// TIA Portal project "N16-1166-5_27082020" (V13)

(* hardware
DEVICE "S71500/ET200MP station_1"  S7-1500 station
   slot 0: "Rail_0"  6ES7 590-1***0-0AA0
   slot 1: "PLC1"  CPU 1513-1 PN  6ES7 513-1AL01-0AB0  V1.8
DEVICE "ET 200SP station_1"  ET 200SP-Station
   slot 0: "Rack_0"  6ES5 710-8MAx1
   slot 0: "pa30"  IM155-6 PN BA  6ES7 155-6AR00-0AN0  V3.2
   slot 1: "DI A11"  DI 8x24VDC ST  6ES7 131-6BF00-0BA0  V1.1
      slot 1: "DI A11"  DI 8x24VDC ST  6ES7 131-6BF00-0BA0
   slot 2: "DI A12"  DI 8x24VDC ST  6ES7 131-6BF00-0BA0  V1.0
      slot 1: "DI A12"  DI 8x24VDC ST  6ES7 131-6BF00-0BA0
   slot 3: "DQ A13"  8DO 24VDC/0,5A ST  6ES7 132-6BF00-0BA0  V1.1
      slot 1: "DQ A13"  DQ 8x24VDC/0.5A ST  6ES7 132-6BF00-0BA0
   slot 4: "CM PtP A14"  CM PtP  6ES7 137-6AA00-0BA0  V1.0
      slot 1: "CM PtP A14"  CM PtP Sub  6ES7 137-6AA00-0BA0
   slot 5: "DI A15"  DI 16x24VDC ST  6ES7 131-6BH00-0BA0  V1.1
      slot 1: "DI A15"  DI 16x24VDC ST  6ES7 131-6BH00-0BA0
   slot 6: "DQ A16"  DQ 16x24VDC/0.5A ST  6ES7 132-6BH00-0BA0  V1.1
      slot 1: "DQ A16"  DQ 16x24VDC/0.5A ST  6ES7 132-6BH00-0BA0
   slot 7: "DI A17"  DI 8x24VDC ST  6ES7 131-6BF00-0BA0  V1.1
      slot 1: "DI A17"  DI 8x24VDC ST  6ES7 131-6BF00-0BA0
   slot 8: "Server module_1"  Server module  6ES7 193-6PA00-0AA0  V1.0
      slot 1: "Server module_1"  Server module  6ES7 193-6PA00-0AA0
   slot 127: "PROFINET BusAdapter CU"  PROFINET Interface  6ES7 193-6AR00-0AA0  V0.0
      slot 1: "Port_1"  6ES7 193-6AR00-0AA0  V0.0
      slot 2: "Port_2"  6ES7 193-6AR00-0AA0  V0.0
DEVICE "ET 200SP station_3"  ET 200SP-Station
   slot 0: "Rack_0"  6ES5 710-8MAx1
   slot 0: "pa60"  IM155-6 PN BA  6ES7 155-6AR00-0AN0  V3.2
   slot 1: "DI 8x24VDC ST_1"  DI 8x24VDC ST  6ES7 131-6BF00-0BA0  V1.1
      slot 1: "DI 8x24VDC ST_1"  DI 8x24VDC ST  6ES7 131-6BF00-0BA0
   slot 2: "DI 8x24VDC ST_2"  DI 8x24VDC ST  6ES7 131-6BF00-0BA0  V1.0
      slot 1: "DI 8x24VDC ST_2"  DI 8x24VDC ST  6ES7 131-6BF00-0BA0
   slot 3: "DI 8x24VDC ST_3"  DI 8x24VDC ST  6ES7 131-6BF00-0BA0  V1.1
      slot 1: "DI 8x24VDC ST_3"  DI 8x24VDC ST  6ES7 131-6BF00-0BA0
   slot 4: "DQ 8x24VDC/0.5A ST_1"  8DO 24VDC/0,5A ST  6ES7 132-6BF00-0BA0  V1.1
      slot 1: "DQ 8x24VDC/0.5A ST_1"  DQ 8x24VDC/0.5A ST  6ES7 132-6BF00-0BA0
   slot 5: "CM PtP_1"  CM PtP  6ES7 137-6AA00-0BA0  V1.0
      slot 1: "CM PtP_1"  CM PtP Sub  6ES7 137-6AA00-0BA0
   slot 6: "DI 16x24VDC ST_1"  DI 16x24VDC ST  6ES7 131-6BH00-0BA0  V1.1
      slot 1: "DI 16x24VDC ST_1"  DI 16x24VDC ST  6ES7 131-6BH00-0BA0
   slot 7: "DQ 16x24VDC/0.5A ST_1"  DQ 16x24VDC/0.5A ST  6ES7 132-6BH00-0BA0  V1.1
      slot 1: "DQ 16x24VDC/0.5A ST_1"  DQ 16x24VDC/0.5A ST  6ES7 132-6BH00-0BA0
   slot 8: "Server module_1"  Server module  6ES7 193-6PA00-0AA0  V1.0
      slot 1: "Server module_1"  Server module  6ES7 193-6PA00-0AA0
   slot 127: "PROFINET BusAdapter CU"  PROFINET Interface  6ES7 193-6AR00-0AA0  V0.0
      slot 1: "Port_1"  6ES7 193-6AR00-0AA0  V0.0
      slot 2: "Port_2"  6ES7 193-6AR00-0AA0  V0.0
DEVICE "HMI_pa30"  KTP700 Basic PN
   slot 0: "HMI"  HMI  6AV2 123-2GB03-0AX0  13.0.1.0
   slot 1: "HMI_RT_2"  KTP700 Basic PN  6AV2 123-2GB03-0AX0  13.0.1.0
   slot 5: "HMI_pa30.IE_CP_1"  PROFINET Interface
      slot 1: "PROFINET Interface_1"  PROFINET Interface
         slot 1: "Port_1"  Port
DEVICE "HMI_pa60"  KTP700 Basic PN
   slot 0: "HMI"  HMI  6AV2 123-2GB03-0AX0  13.0.1.0
   slot 1: "HMI_RT_4"  KTP700 Basic PN  6AV2 123-2GB03-0AX0  13.0.1.0
   slot 5: "HMI_pa60.IE_CP_1"  PROFINET Interface
      slot 1: "PROFINET Interface_1"  PROFINET Interface
         slot 1: "Port_1"  Port
DEVICE "ET 200SP station_4"  ET 200SP-Station
   slot 0: "Rack_0"  6ES5 710-8MAx1
   slot 0: "LightControll"  IM155-6 PN BA  6ES7 155-6AR00-0AN0  V3.2
   slot 1: "DQ 16x24VDC/0.5A ST_1"  DQ 16x24VDC/0.5A ST  6ES7 132-6BH00-0BA0  V1.1
      slot 1: "DQ 16x24VDC/0.5A ST_1"  DQ 16x24VDC/0.5A ST  6ES7 132-6BH00-0BA0
   slot 2: "Server module_1"  Server module  6ES7 193-6PA00-0AA0  V1.0
      slot 1: "Server module_1"  Server module  6ES7 193-6PA00-0AA0
   slot 127: "PROFINET BusAdapter CU"  PROFINET Interface  6ES7 193-6AR00-0AA0  V0.0
      slot 1: "Port_1"  6ES7 193-6AR00-0AA0  V0.0
      slot 2: "Port_2"  6ES7 193-6AR00-0AA0  V0.0
DEVICE "S71500/ET200MP station_2"  S7-1500 station
   slot 0: "Rail_0"  6ES7 590-1***0-0AA0
   slot 2: "CP 1543-1_1"  CP 1543-1  6GK7 543-1AX00-0XE0  V1.1
DEVICE "HMI_PA10B"  KTP700 Basic PN
   slot 0: "HMI"  HMI  6AV2 123-2GB03-0AX0  13.0.1.0
   slot 1: "HMI_RT_5"  KTP700 Basic PN  6AV2 123-2GB03-0AX0  13.0.1.0
   slot 5: "HMI_PA10B.IE_CP_1"  PROFINET Interface
      slot 1: "PROFINET Interface_1"  PROFINET Interface
         slot 1: "Port_1"  Port
DEVICE "ET 200SP station_5"  ET 200SP-Station
   slot 0: "Rack_0"  6ES5 710-8MAx1
   slot 0: "FS"  IM155-6 PN BA  6ES7 155-6AR00-0AN0  V3.2
   slot 1: "DI 8x24VDC ST_1"  DI 8x24VDC ST  6ES7 131-6BF00-0BA0  V1.0
      slot 1: "DI 8x24VDC ST_1"  DI 8x24VDC ST  6ES7 131-6BF00-0BA0
   slot 2: "DI 8x24VDC ST_2"  DI 8x24VDC ST  6ES7 131-6BF00-0BA0  V1.1
      slot 1: "DI 8x24VDC ST_2"  DI 8x24VDC ST  6ES7 131-6BF00-0BA0
   slot 3: "DI 8x24VDC ST_3"  DI 8x24VDC ST  6ES7 131-6BF00-0BA0  V1.1
      slot 1: "DI 8x24VDC ST_3"  DI 8x24VDC ST  6ES7 131-6BF00-0BA0
   slot 4: "DI 8x24VDC ST_4"  DI 8x24VDC ST  6ES7 131-6BF00-0BA0  V1.1
      slot 1: "DI 8x24VDC ST_4"  DI 8x24VDC ST  6ES7 131-6BF00-0BA0
   slot 5: "DI 8x24VDC ST_5"  DI 8x24VDC ST  6ES7 131-6BF00-0BA0  V1.1
      slot 1: "DI 8x24VDC ST_5"  DI 8x24VDC ST  6ES7 131-6BF00-0BA0
   slot 6: "CM PtP_1"  CM PtP  6ES7 137-6AA00-0BA0  V1.0
      slot 1: "CM PtP_1"  CM PtP Sub  6ES7 137-6AA00-0BA0
   slot 7: "DI 16x24VDC ST_1"  DI 16x24VDC ST  6ES7 131-6BH00-0BA0  V1.1
      slot 1: "DI 16x24VDC ST_1"  DI 16x24VDC ST  6ES7 131-6BH00-0BA0
   slot 8: "DQ 16x24VDC/0.5A ST_1"  DQ 16x24VDC/0.5A ST  6ES7 132-6BH00-0BA0  V1.1
      slot 1: "DQ 16x24VDC/0.5A ST_1"  DQ 16x24VDC/0.5A ST  6ES7 132-6BH00-0BA0
   slot 9: "Server module_1"  Server module  6ES7 193-6PA00-0AA0  V1.0
      slot 1: "Server module_1"  Server module  6ES7 193-6PA00-0AA0
   slot 127: "PROFINET BusAdapter CU"  PROFINET Interface  6ES7 193-6AR00-0AA0  V0.0
      slot 1: "Port_1"  6ES7 193-6AR00-0AA0  V0.0
      slot 2: "Port_2"  6ES7 193-6AR00-0AA0  V0.0
DEVICE "ET 200SP station_6"  ET 200SP-Station
   slot 0: "Rack_0"  6ES5 710-8MAx1
   slot 0: "PA10B"  IM155-6 PN BA  6ES7 155-6AR00-0AN0  V3.2
   slot 1: "DI 8x24VDC ST_1"  DI 8x24VDC ST  6ES7 131-6BF00-0BA0  V1.1
      slot 1: "DI 8x24VDC ST_1"  DI 8x24VDC ST  6ES7 131-6BF00-0BA0
   slot 2: "DI 8x24VDC ST_2"  DI 8x24VDC ST  6ES7 131-6BF00-0BA0  V1.0
      slot 1: "DI 8x24VDC ST_2"  DI 8x24VDC ST  6ES7 131-6BF00-0BA0
   slot 3: "DI 16x24VDC ST_1"  DI 16x24VDC ST  6ES7 131-6BH00-0BA0  V1.1
      slot 1: "DI 16x24VDC ST_1"  DI 16x24VDC ST  6ES7 131-6BH00-0BA0
   slot 4: "DQ 16x24VDC/0.5A ST_1"  DQ 16x24VDC/0.5A ST  6ES7 132-6BH00-0BA0  V1.1
      slot 1: "DQ 16x24VDC/0.5A ST_1"  DQ 16x24VDC/0.5A ST  6ES7 132-6BH00-0BA0
   slot 5: "DQ 16x24VDC/0.5A ST_2"  DQ 16x24VDC/0.5A ST  6ES7 132-6BH00-0BA0  V1.0
      slot 1: "DQ 16x24VDC/0.5A ST_2"  DQ 16x24VDC/0.5A ST  6ES7 132-6BH00-0BA0
   slot 6: "CM PtP_1"  CM PtP  6ES7 137-6AA00-0BA0  V1.0
      slot 1: "CM PtP_1"  CM PtP Sub  6ES7 137-6AA00-0BA0
   slot 7: "Server module_1"  Server module  6ES7 193-6PA00-0AA0  V1.0
      slot 1: "Server module_1"  Server module  6ES7 193-6PA00-0AA0
   slot 127: "PROFINET BusAdapter CU"  PROFINET Interface  6ES7 193-6AR00-0AA0  V0.0
      slot 1: "Port_1"  6ES7 193-6AR00-0AA0  V0.0
      slot 2: "Port_2"  6ES7 193-6AR00-0AA0  V0.0
DEVICE "ET 200SP station_7"  ET 200SP-Station
   slot 0: "Rack_0"  6ES5 710-8MAx1
   slot 0: "PA20B"  IM155-6 PN BA  6ES7 155-6AR00-0AN0  V3.2
   slot 1: "DI 8x24VDC ST_1"  DI 8x24VDC ST  6ES7 131-6BF00-0BA0  V1.1
      slot 1: "DI 8x24VDC ST_1"  DI 8x24VDC ST  6ES7 131-6BF00-0BA0
   slot 2: "DI 8x24VDC ST_2"  DI 8x24VDC ST  6ES7 131-6BF00-0BA0  V1.0
      slot 1: "DI 8x24VDC ST_2"  DI 8x24VDC ST  6ES7 131-6BF00-0BA0
   slot 3: "DQ 16x24VDC/0.5A ST_1"  DQ 16x24VDC/0.5A ST  6ES7 132-6BH00-0BA0  V1.1
      slot 1: "DQ 16x24VDC/0.5A ST_1"  DQ 16x24VDC/0.5A ST  6ES7 132-6BH00-0BA0
   slot 4: "Server module_1"  Server module  6ES7 193-6PA00-0AA0  V1.0
      slot 1: "Server module_1"  Server module  6ES7 193-6PA00-0AA0
   slot 127: "PROFINET BusAdapter CU"  PROFINET Interface  6ES7 193-6AR00-0AA0  V0.0
      slot 1: "Port_1"  6ES7 193-6AR00-0AA0  V0.0
      slot 2: "Port_2"  6ES7 193-6AR00-0AA0  V0.0
DEVICE "HMI_1"  KTP700 Basic PN
   slot 0: "HMI"  HMI  6AV2 123-2GB03-0AX0  13.0.1.0
   slot 1: "HMI_RT_7"  KTP700 Basic PN  6AV2 123-2GB03-0AX0  13.0.1.0
   slot 5: "HMI_1.IE_CP_1"  PROFINET Interface
      slot 1: "PROFINET Interface_1"  PROFINET Interface
         slot 1: "Port_1"  Port
*)

// ===== PLC "PLC1"  CPU 1513-1 PN =====

VAR_GLOBAL   // PLC tag table "Default tag table"
   "RPA30R_RoofRotationSensorYL" AT %I12.3 : Bool;
   "RPA30R_RoofRotationSensorYAtOperator" AT %I12.2 : Bool;
   "RPA30R_RoofRotationSensorYR" AT %I12.1 : Bool;
   "RPA30R_RoofRotationSensorYFromOperator" AT %I12.0 : Bool;
   "RPA30R_PositionCylinderSensorUnlockY" AT %I12.4 : Bool;
   "RPA30R_PositionCylinderSensorLockY" AT %I12.5 : Bool;
   "RPA30R_SensorIFMLeftTriggerOut" AT %I12.6 : Bool;
   "RPA30R_SensorIFMLeftReadyOut" AT %I12.7 : Bool;
   "RPA30R_SensorIFMLeftOut" AT %I13.0 : Bool;
   "RPA30R_SensorIFMRightTriggerOut" AT %I13.1 : Bool;
   "RPA30R_SensorIFMRightReadyOut" AT %I13.2 : Bool;
   "RPA30R_SensorIFMRightOut" AT %I13.3 : Bool;
   "RPA30R_PrimerPA10SensorPadLeft" AT %I22.0 : Bool;
   "RPA30R_PrimerPA10SensorPadRight" AT %I22.1 : Bool;
   "RPA30R_PrimerPA10SensorFelt" AT %I22.2 : Bool;
   "RPA30R_PrimerPA30SensorRemover208" AT %I22.3 : Bool;
   "RPA30R_PrimerPA30SensorFeltEmpty" AT %I22.4 : Bool;
   "RPA30R_PrimerPA30ButtonPadIsChanged" AT %I22.5 : Bool;
   "RPA30R_LCDSwitchAutomat_Manual" AT %I22.6 : Bool;
   "RPA30R_LCDButtonStart" AT %I22.7 : Bool;
   "RPA30R_LCDButtonConfirmSignal" AT %I23.0 : Bool;
   "RPA30R_PrimerPA30SensorBottleRemover208" AT %I23.1 : Bool;
   "RPA30R_PrimerPA30SensorBottlePrimer207" AT %I23.4 : Bool;
   "RPA60R_RoofRotationSensorYL" AT %I34.3 : Bool;
   "RPA60R_RoofRotationSensorYAtOperator" AT %I34.2 : Bool;
   "RPA60R_RoofRotationSensorYR" AT %I34.1 : Bool;
   "RPA60R_RoofRotationSensorYFromOperator" AT %I34.0 : Bool;
   "RPA60R_valvePositionSensorUnlockY" AT %I34.4 : Bool;
   "RPA60R_valvePositionSensorLockY" AT %I34.5 : Bool;
   "RPA60R_SenzorLoaderPresenceLeft581" AT %I34.6 : Bool;
   "RPA60R_SenzorLoaderPresenceRear581" AT %I34.7 : Bool;
   "RPA60R_SenzorLoaderPresenceRight581" AT %I35.0 : Bool;
   "RPA60R_SenzorLoaderPresenceLeft582" AT %I35.1 : Bool;
   "RPA60R_SenzorLoaderPresenceRear582" AT %I35.2 : Bool;
   "RPA60R_SenzorLoaderPresenceRight582" AT %I35.3 : Bool;
   "RPA60R_SenzorSealPresenceLeft581" AT %I35.4 : Bool;
   "RPA60R_SenzorSealPresenceRear581" AT %I35.5 : Bool;
   "RPA60R_SenzorSealPresenceRight581" AT %I35.6 : Bool;
   "RPA60R_SenzorSealPresenceLeft582" AT %I35.7 : Bool;
   "RPA60R_SenzorSealPresenceRear582" AT %I36.0 : Bool;
   "RPA60R_SenzorSealPresenceRight582" AT %I36.1 : Bool;
   "RPA60R_SenzorVacuum" AT %I36.2 : Bool;
   "RPA60R_LCDSwitchAutomat_Manual" AT %I45.0 : Bool;
   "RPA60R_LCDButtonStart" AT %I45.1 : Bool;
   "RPA60R_LCDButtonConfirmSignal" AT %I45.2 : Bool;
   "RPA60R_SenzorRoller" AT %I36.3 : Bool;
   "RPA20B_belt_position_sensor" AT %I66.0 : Bool;
   "RPA20B_blend_presence_sensor_1" AT %I66.1 : Bool;
   "RPA20B_blend_presence_sensor_2" AT %I66.2 : Bool;
   "RPA20B_drawer_position_sensor" AT %I66.3 : Bool;
   "RPA20B_drawer_lock_sensor" AT %I66.4 : Bool;
   "RPA20B_drawer_unlock_sensor" AT %I66.5 : Bool;
   "RPA20B_ES_feedback" AT %I66.6 : Bool;
   "RPA20B_lock_door_feedback" AT %I66.7 : Bool;
   "RPA20B_manual_UP" AT %I67.0 : Bool;
   "RPA20B_manual_DOWN" AT %I67.1 : Bool;
   "RPA20B_manual_move" AT %I67.2 : Bool;
   "RPA20B_unlock_button" AT %I67.3 : Bool;
   "RPA20B_Camera_Test_Ok" AT %I67.4 : Bool;
   "ib_FS_sensor_bottle_1" AT %I47.0 : Bool;
   "ib_FS_sensor_bottle_2" AT %I47.1 : Bool;
   "ib_FS_sensor_bottle_3" AT %I47.2 : Bool;
   "ib_FS_sensor_bottle_4" AT %I47.3 : Bool;
   "ib_FS_sensor_bottle_5" AT %I47.4 : Bool;
   "ib_FS_mixer_1_presence_sensor_1" AT %I47.5 : Bool;
   "ib_FS_mixer_1_presence_sensor_2" AT %I47.6 : Bool;
   "ib_FS_mixer_2_presence_sensor_1" AT %I47.7 : Bool;
   "ib_FS_mixer_2_presence_sensor_2" AT %I48.0 : Bool;
   "ib_FS_mixer_1_door_1_is_close" AT %I48.1 : Bool;
   "ib_FS_mixer_1_door_2_is_close" AT %I48.2 : Bool;
   "ib_FS_mixer_2_door_1_is_close" AT %I48.3 : Bool;
   "ib_FS_mixer_2_door_2_is_close" AT %I48.4 : Bool;
   "ib_FS_funnel_1_position_sensor_UP" AT %I49.0 : Bool;
   "ib_FS_funnel_1_position_sensor_DOWN" AT %I49.1 : Bool;
   "ib_FS_funnel_2_position_sensor_UP" AT %I49.2 : Bool;
   "ib_FS_funnel_2_position_sensor_DOWN" AT %I49.3 : Bool;
   "ib_FS_funnel_3_position_sensor_UP" AT %I49.4 : Bool;
   "ib_FS_funnel_3_position_sensor_DOWN" AT %I49.5 : Bool;
   "ib_FS_funnel_4_position_sensor_UP" AT %I49.6 : Bool;
   "ib_FS_funnel_4_position_sensor_DOWN" AT %I49.7 : Bool;
   "ib_FS_funnel_5_position_sensor_UP" AT %I50.0 : Bool;
   "ib_FS_funnel_5_position_sensor_DOWN" AT %I50.1 : Bool;
   "ib_FS_mixer_1_door_1_is_unlock" AT %I50.2 : Bool;
   "ib_FS_mixer_1_door_1_is_lock" AT %I50.3 : Bool;
   "ib_FS_mixer_1_door_2_is_unlock" AT %I50.4 : Bool;
   "ib_FS_mixer_1_door_2_is_lock" AT %I50.5 : Bool;
   "ib_FS_mixer_2_door_1_is_unlock" AT %I50.6 : Bool;
   "ib_FS_mixer_2_door_1_is_lock" AT %I50.7 : Bool;
   "ib_FS_mixer_2_door_2_is_unlock" AT %I51.0 : Bool;
   "ib_FS_mixer_2_door_2_is_lock" AT %I51.1 : Bool;
   "ib_FS_LCD_switch_automat_manual" AT %I61.0 : Bool;
   "ib_FS_LCD_button_start" AT %I61.1 : Bool;
   "ib_FS_LCD_button_confirm" AT %I61.2 : Bool;
   "RPA10B_home_position_horizontal_carriage_sensor" AT %I52.0 : Bool;
   "RPA10B_end_position_horizontal_carriage_sensor" AT %I52.1 : Bool;
   "RPA10B_home_position_idler_carriage_sensor" AT %I52.2 : Bool;
   "RPA10B_end_position_idler_carriage_sensor" AT %I52.3 : Bool;
   "RPA10B_code_position_1" AT %I52.4 : Bool;
   "RPA10B_code_position_2" AT %I52.5 : Bool;
   "RPA10B_idler_presence_sensor" AT %I52.6 : Bool;
   "RPA10B_vacuum_sensor" AT %I52.7 : Bool;
   "RPA10B_lock_sensor" AT %I63.1 : Bool;
   "RPA10B_unlock_sensor" AT %I63.2 : Bool;
   "RPA10B_blend_1_vacuum_fix_sensor" AT %I63.3 : Bool;
   "RPA10B_blend_2_vacuum_fix_sensor" AT %I63.4 : Bool;
   "RPA10B_LCD_switch_manual_automat" AT %I64.0 : Bool;
   "RPA10B_LCD_button_start" AT %I64.1 : Bool;
   "RPA10B_LCD_button_confirm" AT %I64.2 : Bool;
   "RPA10B_primerbox_pad_sensor_left" AT %I64.3 : Bool;
   "RPA10B_primerbox_pad_sensor_right" AT %I64.4 : Bool;
   "RPA10B_primerbox_felt_sensor" AT %I64.5 : Bool;
   "RPA10B_primerbox_felt_presence_sensor" AT %I64.6 : Bool;
   "RPA10B_primerbox_button_PAD_IS_CHANGED" AT %I64.7 : Bool;
   "RPA10B_primerbox_bottle_1" AT %I65.0 : Bool;
   "RPA10B_primerbox_bottle_2" AT %I65.1 : Bool;
   "RPA10B_EJ_1_vacuum_sensor" AT %I65.2 : Bool;
   "RPA10B_EJ_2_vacuum_sensor" AT %I65.3 : Bool;
   "RPA10B_universal_button_1" AT %I65.4 : Bool;
   "RPA10B_universal_button_2" AT %I65.5 : Bool;
   "ib_FS_mixer_3_bottle_pressence" AT %I48.5 : Bool;
   "ib_FS_mixer_3_door_position" AT %I48.6 : Bool;
   "RPA30_keyence_right_2" AT %I76.1 : Bool;
   "RPA30_keyence_right_1" AT %I76.0 : Bool;
   "RPA30_keyence_middle_1" AT %I13.6 : Bool;
   "RPA30_keyence_middle_2" AT %I13.7 : Bool;
   "RPA30_keyence_left_1" AT %I13.4 : Bool;
   "RPA30_keyence_left_2" AT %I13.5 : Bool;
   "RPA60R_LH_CAM" AT %I36.6 : Bool;
   "RPA60R_RH_CAM" AT %I36.4 : Bool;
   "RPA10B_Left_Hand_Detection" AT %I63.6 : Bool;
   "RPA10B_Right_Hand_Detection" AT %I63.7 : Bool;
   "RPA20B_Camera_Start_Test" AT %I67.5 : Bool;
   "RPA60R_CAM_START_TEST" AT %I46.4 : Bool;
   "RPA60R_LHI_CAM" AT %I46.2 : Bool;
   "RPA60R_RHI_CAM" AT %I46.0 : Bool;
   "RPA20B_Product_Present_On_Top_Level" AT %I67.6 : Bool;
   "RPA30R_ValveCylinderYLock" AT %Q5.0 : Bool;
   "RPA30R_SensorIFMLeftTrigger" AT %Q5.2 : Bool;
   "RPA30R_SensorIFMLeft_Input_1" AT %Q5.3 : Bool;
   "RPA30R_SensorIFMLeft_Input_2" AT %Q5.4 : Bool;
   "RPA30R_SensorIFMRightTrigger" AT %Q5.5 : Bool;
   "RPA30R_SensorIFMRight_Input_1" AT %Q5.6 : Bool;
   "RPA30R_SensorIFMRight_Input_2" AT %Q5.7 : Bool;
   "RPA30R_Beacon_1_LCDPanelGreen" AT %Q6.0 : Bool;
   "RPA30R_Beacon_1_LCDPanelOrange" AT %Q6.1 : Bool;
   "RPA30R_Beacon_1_LCDPanelRed" AT %Q6.2 : Bool;
   "RPA30R_Beacon_1_LCDPanelSiren" AT %Q6.3 : Bool;
   "RPA30R_Beacon_2_PrimerBoxGreen" AT %Q6.4 : Bool;
   "RPA30R_Beacon_2_PrimerBoxOrange" AT %Q6.5 : Bool;
   "RPA30R_Beacon_2_PrimerBoxRed" AT %Q6.6 : Bool;
   "RPA30R_Beacon_2_PrimerBoxSiren" AT %Q6.7 : Bool;
   "RPA30R_PrimerPA30GreenReady" AT %Q7.0 : Bool;
   "RPA30R_PrimerPA30GreenFelt" AT %Q7.1 : Bool;
   "RPA30R_PrimerPA30GreenRemover208" AT %Q7.2 : Bool;
   "RPA30R_PrimerPA30GreenPrimer207" AT %Q7.3 : Bool;
   "RPA30R_PrimerPA30RedNotReady" AT %Q7.4 : Bool;
   "RPA30R_PrimerPA30RedChangePad" AT %Q7.5 : Bool;
   "RPA30R_LEDGreenSart" AT %Q7.6 : Bool;
   "RPA30R_LedBlueConfirm" AT %Q7.7 : Bool;
   "RPA60R_ValveCylinderYLock" AT %Q10.0 : Bool;
   "RPA60R_Beacon_1_LCDPanelGreen" AT %Q11.0 : Bool;
   "RPA60R_Beacon_1_LCDPanelOrange" AT %Q11.1 : Bool;
   "RPA60R_Beacon_1_LCDPanelRed" AT %Q11.2 : Bool;
   "RPA60R_Beacon_1_LCDPanelSiren" AT %Q11.3 : Bool;
   "RPA60R_LEDGreenSart" AT %Q11.4 : Bool;
   "RPA60R_LedBlueConfirm" AT %Q11.5 : Bool;
   "RPA10R_light" AT %Q13.0 : Bool;
   "RPA30R_light" AT %Q13.1 : Bool;
   "RPA50R_light" AT %Q13.2 : Bool;
   "RPA60R_light" AT %Q13.3 : Bool;
   "RPA60R_VacuumSwitch" AT %Q10.1 : Bool;
   "RPA60R_LEDRoller" AT %Q11.6 : Bool;
   "RPA20B_open_drawer" AT %Q21.0 : Bool;
   "RPA20B_open_door_LED_green" AT %Q21.1 : Bool;
   "RPA20B_button_back_LED_1" AT %Q21.2 : Bool;
   "RPA20B_button_back_LED_2" AT %Q21.3 : Bool;
   "RPA20B_valve_close_drawer" AT %Q21.4 : Bool;
   "RPA20B_valve_open_drawer" AT %Q21.5 : Bool;
   "ob_FS_LCD_beacon_green" AT %Q15.0 : Bool;
   "ob_FS_LCD_beacon_orange" AT %Q15.1 : Bool;
   "ob_FS_LCD_beacon_red" AT %Q15.2 : Bool;
   "ob_FS_LCD_beacon_siren" AT %Q15.3 : Bool;
   "ob_FS_LCD_start_button_LED_green" AT %Q15.4 : Bool;
   "ob_FS_LCD_confirm_button_LED_blue" AT %Q15.5 : Bool;
   "ob_FS_move_UP_funel_1" AT %Q15.6 : Bool;
   "ob_FS_move_UP_funel_2" AT %Q15.7 : Bool;
   "ob_FS_move_UP_funel_3" AT %Q16.0 : Bool;
   "ob_FS_move_UP_funel_4" AT %Q16.1 : Bool;
   "ob_FS_move_UP_funel_5" AT %Q16.2 : Bool;
   "ob_FS_mixer_1_door_1_lock" AT %Q16.3 : Bool;
   "ob_FS_mixer_1_door_2_lock" AT %Q16.4 : Bool;
   "ob_FS_mixer_2_door_1_lock" AT %Q16.5 : Bool;
   "ob_FS_mixer_2_door_2_lock" AT %Q16.6 : Bool;
   "RPA10B_LCD_beacon_green" AT %Q17.0 : Bool;
   "RPA10B_LCD_beacon_orange" AT %Q17.1 : Bool;
   "RPA10B_LCD_beacon_red" AT %Q17.2 : Bool;
   "RPA10B_LCD_beacon_siren" AT %Q17.3 : Bool;
   "RPA10B_primerbox_beacon_green" AT %Q17.4 : Bool;
   "RPA10B_primerbox_beacon_orange" AT %Q17.5 : Bool;
   "RPA10B_primerbox_beacon_red" AT %Q17.6 : Bool;
   "RPA10B_primerbox_beacon_siren" AT %Q17.7 : Bool;
   "RPA10B_primerbox_LED_green_ready" AT %Q18.0 : Bool;
   "RPA10B_primerbox_LED_green_felt" AT %Q18.1 : Bool;
   "RPA10B_primerbox_LED_green_bottle_1" AT %Q18.2 : Bool;
   "RPA10B_primerbox_LED_green_bottle_2" AT %Q18.3 : Bool;
   "RPA10B_primerbox_LED_red_NOT_READY" AT %Q18.4 : Bool;
   "RPA10B_primerbox_LED_orange_change_pad" AT %Q18.5 : Bool;
   "RPA10B_LCD_LED_green_start_button" AT %Q18.6 : Bool;
   "RPA10B_LCD_LED_blue_confirm_button" AT %Q18.7 : Bool;
   "RPA10B_vavle_aretation_unlock" AT %Q19.0 : Bool;
   "RPA10B_vavle_aretation_lock" AT %Q19.1 : Bool;
   "RPA10B_vavle_seal_idler_unlock" AT %Q19.2 : Bool;
   "RPA10B_vavle_seal_idler_lock" AT %Q19.3 : Bool;
   "RPA10B_EJ_1_vacuum_control" AT %Q19.4 : Bool;
   "RPA10B_EJ_1_eject" AT %Q19.5 : Bool;
   "RPA10B_EJ_2_vacuum_control" AT %Q19.6 : Bool;
   "RPA10B_EJ_2_eject" AT %Q19.7 : Bool;
   "RPA10B_light" AT %Q13.4 : Bool;
   "RPA10B_vacuum_cleaner_switch" AT %Q13.5 : Bool;
   "RPA20_motor_up" AT %Q13.7 : Bool;
   "RPA20B_motor_down" AT %Q14.0 : Bool;
   "ob_FS_mixer_3_door_lock" AT %Q16.7 : Bool;
   "RPA20B_Camera_Trigger" AT %Q22.0 : Bool;
   "RPA20B_Camera_TrafficLight_Green" AT %Q22.1 : Bool;
   "RPA20B_Camera_TrafficLight_Yellow" AT %Q22.2 : Bool;
   "RPA20B_Camera_TrafficLight_Red" AT %Q22.3 : Bool;
   "Clock_Byte" AT %MB0 : Byte;
   "Clock_10Hz" AT %M0.0 : Bool;
   "Clock_5Hz" AT %M0.1 : Bool;
   "Clock_2.5Hz" AT %M0.2 : Bool;
   "Clock_2Hz" AT %M0.3 : Bool;
   "Clock_1.25Hz" AT %M0.4 : Bool;
   "Clock_1Hz" AT %M0.5 : Bool;
   "Clock_0.625Hz" AT %M0.6 : Bool;
   "Clock_0.5Hz" AT %M0.7 : Bool;
   "Tag_1" AT %M10.0 : Bool;
   "RPA60R_CAM_T_START" AT %M100.0 : Bool;
   "RPA60R_CAM_T_RELEASE" AT %M100.1 : Bool;
   "RPA10B_Bottle_1_Left_Side_Applied" AT %M15.0 : Bool;
   "RPA10B_Bottle_1_Right_Side_Applied" AT %M15.1 : Bool;
   "RPA10B_B1_Bottle_1_Applied" AT %M15.2 : Bool;
   "RPA10B_B2_Bottle_1_Applied" AT %M15.3 : Bool;
   "RPA10B_Wipe_Sealing_Surface_Left_Side" AT %M16.0 : Bool;
   "RPA10B_Wipe_Sealing_Surface_Right_Side" AT %M16.1 : Bool;
   "RPA10B_Apply_Activator_Left_Side" AT %M17.0 : Bool;
   "RPA10B_Apply_Activator_Right_Side" AT %M17.1 : Bool;
   "RPA20B_Camera_Result_OK" AT %M20.0 : Bool;
   "RPA20B_Camera_Result_NOK" AT %M20.1 : Bool;
   "RPA_60R_CAM_TEST_1_DONE" AT %M100.2 : Bool;
   "RPA_60R_CAM_TEST_2_DONE" AT %M100.3 : Bool;
END_VAR

VAR_GLOBAL CONSTANT   // PLC tag table "Default tag table"
   "RPA20B_push_start_button" : Int := 0;
   "RPA20B_wait_to_deactivate_belt_sensor" : Int := 1;
   "RPA20B_wait_to_activate_belt_sensor" : Int := 2;
   "RPA20B_wait_to_deactivate_start_button" : Int := 3;
   "RPA20B_wait_for_deactivate_open_button" : Int := 4;
   "RPA20B_wait_to_push_open_button" : Int := 0;
   "RPA20B_open_drawer_state" : Int := 6;
   "RPA20B_wait_to_push_close_button" : Int := 7;
   "RPA20B_close_drawer_state" : Int := 8;
   "RPA20B_is_blend_release" : Int := 9;
   "RPA20B_end_operation" : Int := 10;
   "RPA10B_go_to_home_position" : UInt := 0;
   "RPA10B_hmi_go_to_home_position" : Byte := 0;
   "RPA10B_hmi_scan_covers" : Byte := 1;
   "RPA10B_hmi_place_right_cover" : Byte := 2;
   "RPA10B_hmi_place_left_cover" : Byte := 3;
   "RPA10B_place_left_cover" : UInt := 1;
   "RPA10B_place_right_cover" : UInt := 2;
   "RPA10B_take_bottle_1" : UInt := 3;
   "RPA10B_hmi_take_bottle_of_activator" : Byte := 4;
   "RPA10B_scan_bottle_1" : UInt := 4;
   "RPA10B_hmi_scan_bottle" : Byte := 9;
   "RPA10B_change_pad_bottle_1" : UInt := 5;
   "RPA10B_hmi_change_pad" : Byte := 5;
   "RPA10B_hmi_apply_activator" : Byte := 6;
   "RPA10B_apply_bottle" : UInt := 6;
   "RPA10B_take_feld" : UInt := 8;
   "RPA10B_put_back_bottle_1" : UInt := 7;
   "RPA10B_hmi_take_feld" : Byte := 7;
   "RPA10B_hmi_whipe_off" : Byte := 8;
   "RPA10B_whipe_off" : UInt := 9;
   "RPA10B_hmi_stick_sealing_on_right_cover" : Byte := 12;
   "RPA10B_stick_sealing_on_cover_1" : UInt := 10;
   "RPA10B_hmi_press_universal_button_to_use_roller" : Byte := 11;
   "RPA10B_press_universal_button_to_use_roller" : UInt := 12;
   "RPA10B_vacuum_cleaner_cover_1_off" : UInt := 11;
   "RPA10B_stick_sealing_on_cover_2" : UInt := 13;
   "RPA10B_vacuum_cleaner_cover_2_off" : UInt := 14;
   "RPA10B_roller_move_1" : UInt := 15;
   "RPA10B_roller_move_2" : UInt := 16;
   "RPA20B_blend_expiration_checking" : Int := 11;
   "RPA10B_move_roller_to_second_position" : UInt := 17;
   "RPA10B_unlock_axis" : UInt := 18;
   "RPA10B_hmi_Press_button_to_release_left_couver" : Byte := 14;
   "RPA10B_hmi_turn_fixture_to_left_cover" : Byte := 17;
   "RPA10B_rotate_to_left_cover" : UInt := 19;
   "RPA10B_rotate_to_right_cover" : UInt := 20;
   "RPA10B_interposition_1" : UInt := 21;
   "RPA10B_hmi_turn_fixture_to_right_cover" : Byte := 16;
   "RPA10B_take_bottle_2" : UInt := 22;
   "RPA10B_scan_bottle_2" : UInt := 23;
   "RPA10B_change_pad_bottle_2" : UInt := 24;
   "RPA10B_put_back_bottle_2" : UInt := 25;
   "RPA10B_hmi_press_spacers_with_the_tool" : Byte := 13;
   "RPA10B_press_spacers_with_the_tool" : UInt := 26;
   "RPA10B_spacer_usage_dalay" : UInt := 27;
   "RPA10B_put_spacer_back" : UInt := 28;
   "RPA10B_interposition_2" : UInt := 29;
   "RPA10B_interposition_3" : UInt := 30;
   "RPA10B_interposition_4" : UInt := 31;
   "RPA10B_go_home_position_to_finish" : UInt := 32;
   "RPA10B_whipe_off_vacuum_cleaner_off" : UInt := 33;
   "RPA10B_press_button_to_release_right_cover" : UInt := 34;
   "RPA10B_eject_left_cover" : UInt := 35;
   "RPA10B_wait_to_eject_button_release" : UInt := 36;
   "RPA10B_eject_right_cover" : UInt := 40;
   "RPA10B_hmi_press_button_to_release_right_couver" : Byte := 15;
   "RPA10B_press_button_to_release_left_cover" : UInt := 37;
   "RPA10B_end_of_cyclus" : UInt := 38;
   "RPA10B_cyclus_finished_OK" : Byte := 18;
   "RPA10B_reset_cyclus" : UInt := 50;
   "RPA30_reset_cyclus" : UInt := 90;   // společné pro všechny mody
   "RPA30_go_to_home_position" : UInt := 0;   // společné pro všechny mody
   "RPA60_go_to_home_position" : UInt := 0;
   "RPA60_reset_cyclus" : UInt := 90;
   "RPA10B_active_RPA20B" : UInt := 51;
   "RPA10B_hmi_active_carring_buffer" : Byte := 19;
   "RPA10B_hmi_stick_sealing_on_left_cover" : Byte := 20;
   "RPA10B_switch_on_caring_buffer" : UInt := 52;
   "RPA10B_carring_buffer_full" : UInt := 53;
   "RPA60_check_hardware_configuration" : UInt := 1;
   "RPA60_bad_hardware_configuration" : UInt := 2;
   "RPA60_scan_frame" : UInt := 3;
   "RPA60_bad_frame_code" : UInt := 4;
   "RPA60_bad_frame_hardware_configuration" : UInt := 5;
   "RPA60_unlock_axis" : UInt := 6;
   "RPA60_turn_to_side_2" : UInt := 7;
   "RPA60_end_of_cyclus" : UInt := 8;
   "RPA60_turn_to_side_3" : UInt := 9;
   "RPA60_turn_to_side_4" : UInt := 10;
   "RPA60_check_seals_presence" : UInt := 11;
   "RPA60_seals_presence_error" : UInt := 12;
   "RPA60_print_label" : UInt := 13;
   "RPA60_scan_printed_label" : UInt := 14;
   "RPA60_print_label_agin" : UInt := 15;
   "RPA60_put_sealing_in_the_ficture" : UInt := 16;
   "RPA60_press_sealing_with_roller" : UInt := 17;
   "RPA60_put_roller_to_home_position" : UInt := 18;
   "RPA60_unlock_axis_after_cyclus" : UInt := 19;
   "RPA60_return_to_home_position" : UInt := 20;
   "RPA60_hmi_go_to_home_position" : Byte := 0;
   "RPA60_hmi_scan_frame" : Byte := 3;
   "RPA60_hmi_turn_frame_clockwise" : Byte := 7;
   "RPA60_hmi_put_sealing_in_the_ficture" : Byte := 8;
   "RPA60_hmi_press_sealing_with_roller" : Byte := 9;
   "RPA60_hmi_put_roller_to_home_position" : Byte := 11;
   "RPA60_hmi_seals_pressence_testing" : Byte := 23;
   "RPA60_hmi_seals_missing" : Byte := 24;
   "RPA60_hmi_scan_printed_label" : Byte := 26;
   "RPA60_hmi_label_is_wrong" : Byte := 27;
   "RPA60_hmi_cyclus_finished_ok" : Byte := 28;
   "RPA30_hmi_go_to_home_position" : Byte := 0;
   "RPA30_scan_frame" : UInt := 1;
   "RPA30_hmi_scan_frame" : Byte := 1;
   "RPA30_frame_not_exists_in_db" : UInt := 2;
   "RPA30_unlock_axis" : UInt := 3;
   "RPA30_turn_frame_on_side_2" : UInt := 4;
   "RPA30_hmi_turn_frame_clockwise" : Byte := 4;
   "RPA30_take_felt" : UInt := 5;
   "RPA30_hmi_take_felt" : Byte := 19;
   "RPA30_on_felt_apply_remover" : UInt := 6;
   "RPA30_hmi_on_felt_apply_remover" : Byte := 20;
   "RPA30_hmi_apply_remover_on_5_points" : Byte := 21;
   "RPA30_ifm_check_on_side_2" : UInt := 7;
   "RPA30_turn_frame_on_side_3" : UInt := 8;
   "RPA30_hmi_turn_frame_counterclockwise" : Byte := 22;
   "RPA30_hmi_apply_primer_on_5_points" : Byte := 9;
   "RPA30_ifm_check_side_3" : UInt := 9;
   "RPA30_turn_frame_to_side_4" : UInt := 10;
   "RPA30_ifm_check_side_4" : UInt := 11;
   "RPA30_take_bottle_of_primer" : UInt := 12;
   "RPA30_scan_bottle_of_primer" : UInt := 13;
   "RPA30_hmi_scan_primer_bottle" : Byte := 6;
   "RPA30_hmi_take_bottle_of_primer" : Byte := 5;
   "RPA30_hmi_change_pad" : Byte := 7;
   "RPA30_change_pad" : UInt := 14;
   "RPA30_put_primer_bottle_back" : UInt := 15;
   "RPA30_hmi_put_primer_bottle_back" : Byte := 16;
   "RPA30_end_of_cylus" : UInt := 17;
   "RPA30_hmi_end_of_cyclus" : Byte := 18;
   "RPA30_hmi_wipe_off" : Byte := 23;
   "RPA30_clean_scaner_receave_buffer" : UInt := 18;
   "RPA30_send_frame_info_to_db" : UInt := 19;
   "RPA30_check_frame_expiration" : UInt := 20;
   "RPA30_check_frame_configuration" : UInt := 21;
   "RPA30_bad_frame_configuration" : UInt := 22;
   "RPA30_frame_expiration_min" : UInt := 23;
   "RPA30_write_bottle_1_to_db" : UInt := 24;
   "RPA30_write_bottle_2_to_db" : UInt := 25;
   "RPA30_write_time_to_db" : UInt := 26;
   "RPA30_frame_expiration_max" : UInt := 27;
   "RPA30_check_station_frame_process" : UInt := 28;
   "RPA30_station_frame_process_error" : UInt := 29;
   "RPA60_check_frame_configuration" : UInt := 21;
   "RPA60_bad_frame_configuration" : UInt := 22;
   "RPA60_frame_not_exists_in_db" : UInt := 23;
   "RPA60_check_frame_expiration_pa10" : UInt := 24;
   "RPA60_check_frame_expiration_pa30" : UInt := 25;
   "RPA60_frame_max_expiration_error" : UInt := 26;
   "RPA60_frame_min_expiration_error" : UInt := 27;
   "RPA60_check_station_process" : UInt := 30;
   "RPA60_station_proccess_error" : UInt := 31;
   "RPA60_check_pre_station_process" : UInt := 32;
   "RPA60_pre_station_process_error" : UInt := 33;
   "RPA60_write_data_to_database" : UInt := 34;
   "RPA60_get_order" : UInt := 35;
   "RPA60_get_frame_record" : UInt := 36;
   "RPA60_remove_record" : UInt := 37;
   "RPA10B_scan_left_cover" : UInt := 54;
   "RPA10B_hmi_scan_left_cover" : Byte := 21;
   "RPA10B_hmi_scan_right_cover" : Byte := 22;
   "RPA10B_scan_right_cover" : UInt := 55;
   "RPA20B_get_blend_time" : Int := 12;
   "RPA10B_write_right_cover_to_db" : UInt := 56;
   "RPA10B_write_left_cover_to_db" : UInt := 57;
   "RPA10B_move_roller_to_home_position" : UInt := 58;
   "RPA10B_hmi_move_roller_to_home_position" : Byte := 23;
   "RPA30_hmi_scan_remover_bottle" : Byte := 24;
   "RPA10B_hmi_apply_activator_on_surface" : Byte := 24;
   "RPA60_recheck_seals" : UInt := 38;
   "RPA60_hmi_check_agin" : Byte := 29;
   "FS_do_nothing" : UInt := 0;
   "FS_reset_cyclus" : UInt := 1;
   "FS_hmi_choose_chemical" : Byte := 0;
   "FS_print_sp_bottle_label_ac" : UInt := 2;
   "RPA10B_hmi_move_roller_to_left_cover" : Byte := 25;
   "FS_print_sp_bottle_label_pr" : UInt := 3;
   "FS_hmi_choose_the_operation" : Byte := 1;
   "FS_scan_sp_label_ac" : UInt := 5;
   "FS_hmi_scan_printed_label" : Byte := 2;
   "FS_check_befor_shaking" : UInt := 6;
   "FS_hmi_scan_suplier_bottle" : Byte := 5;
   "FS_shake_bottle" : UInt := 7;
   "FS_close_shaker_door" : UInt := 8;
   "FS_hmi_close_shaker_door" : Byte := 6;
   "FS_hmi_put_bottle_tp_shaker" : Byte := 3;
   "RPA10B_check_cover_revork" : UInt := 60;
   "RPA30_hmi_check_frame_rework" : UInt := 30;
   "RPA30_write_frame_to_database" : UInt := 31;
   "RPA30_rework_increase" : UInt := 32;
   "RPA30_three_times_and_stop" : UInt := 33;
   "RPA60_increase_rework" : UInt := 100;
   "RPA60_three_times_and_stop" : UInt := 110;
   "RPA30_update_produce_time" : UInt := 34;
   "RPA60_update_process_time" : UInt := 120;
   "RPA30_set_frame_cyclus_to_default" : UInt := 35;
   "RPA30_update_frame_cyclus_state" : UInt := 36;
   "RPA60_check_pre_station_cyclus_complete" : UInt := 130;
   "RPA60_set_frame_cyclus_to_default" : UInt := 140;
   "RPA60_update_frame_cyclus_state" : UInt := 150;
   "RPA60_pre_station_cyclus_complete_error" : UInt := 160;
   "RPA60_generate_csv" : UInt := 170;
   "RPA60_camera_signal_missing" : UInt := 39;
   "RPA60_hmi_RH_camera_filtz_missing" : Byte := 40;
   "RPA60_hmi_LH_camera_filtz_missing" : Byte := 41;
   "RPA10B_hmi_second_whipe_off" : Byte := 70;
   "RPA60_hmi_camera_start_test" : Byte := 42;
END_VAR

TYPE "bottleDataStructure"
VERSION : 0.1
   STRUCT
      BareCode : String;
      "Author" : String;
      filling_date : Date_And_Time;
   END_STRUCT;
END_TYPE

TYPE "frameDataStruct_B"
VERSION : 0.1
   STRUCT
      frameCode : String;
      PA10_dateTime : DTL;
      codeBottle1 : String;
      codeBottle2 : String;
      codeBottle3 : String;
      codeBottle4 : String;
      PA30_dateTime : DTL;
      codeBottle5 : String;
      codeBottle6 : String;
      PA50_dateTime : DTL;
      PA60_dateTime : DTL;
      frameOrder : Int;
      frame_type : Byte;
   END_STRUCT;
END_TYPE

TYPE "instruction_data_list"
VERSION : 0.1
   STRUCT
      list : Array[0..128] of String;
   END_STRUCT;
END_TYPE

TYPE "blendDatatype"
VERSION : 0.1
   STRUCT
      timeExpiration : Int;
   END_STRUCT;
END_TYPE

TYPE "shakerStruct"
VERSION : 0.1
   STRUCT
      chemics : UInt;
      shakeTimeStart : DTL;
      shakerBottleSensor : Bool;
   END_STRUCT;
END_TYPE

TYPE "expirationStruct"
VERSION : 0.1
   STRUCT
      ID : UInt;
      chemical : String;
      shakingEndTime : DTL;
   END_STRUCT;
END_TYPE

TYPE "frameDataStruct_A"
VERSION : 0.1
   STRUCT
      PA30_dateTime : DTL;
      frameCode : String;
      codeBottle1 : String;
      codeBottle2 : String;
      PA60_dateTime : DTL;
      frameOrder : Int;
      frame_type : Byte;
   END_STRUCT;
END_TYPE

TYPE "tcp_data_item"
VERSION : 0.1
   STRUCT
      tcp_item : Array[0..1023] of Char;
   END_STRUCT;
END_TYPE

TYPE "tcp_data_structure"
VERSION : 0.1
   STRUCT
      input_buffer : Array[0..5] of "tcp_data_item";
      output_buffer : Array[0..5] of "tcp_data_item";
      transaction_done : Array[0..5] of Bool;
      size_out : Array[0..5] of UInt;
   END_STRUCT;
END_TYPE

TYPE "fs_data_struct"
VERSION : 0.1
   STRUCT
      funel : Array[0..4] of Bool;
   END_STRUCT;
END_TYPE

DATA_BLOCK "DB_chemical_code"   // DB1
{ S7_Optimized_Access := 'FALSE' }
VERSION : 0.1
   VAR RETAIN
      Supplier_bottle_code_Primer_DV954V1 : String;
      Supplier_bottle_code_Activator_DW646 : String;
      Supplier_bottle_code_Remover_SIKA_208 : String;
      Supplier_bottle_code_Primer_SIKA_207 : String;
      Supplier_bottle_code_Activator_SIKA_110 : String;
      Application_bottle_code_Primer_DV954V1 : String;
      Application_bottle_code_Activator_DW646 : String;
      Application_bottle_code_Remover_SIKA_208 : String;
      Application_bottle_code_Primer_SIKA_207 : String;
      Application_bottle_code_Activator_SIKA_110 : String;
   END_VAR
BEGIN
END_DATA_BLOCK

DATA_BLOCK "filling_station_main_DB"   // DB2
{ S7_Optimized_Access := 'FALSE' }
VERSION : 0.1
// stored: InstanceOfName filling_station_main
"filling_station_main"
BEGIN
END_DATA_BLOCK

DATA_BLOCK "activator_wipe_off"   // DB3
{ S7_Optimized_Access := 'FALSE' }
VERSION : 0.1
   VAR
      left_blend_activator_wipe_off : Int;
      right_blend_activator_wipe_off : Int;
      wipe_off_number_settings : Int;
   END_VAR
BEGIN
END_DATA_BLOCK

DATA_BLOCK "RPA30_DataBlock"   // DB4
{ S7_Optimized_Access := 'FALSE' }
VERSION : 0.1
   VAR
      RPA30_FrameDateTime : DTL;
      RPA30_actualCodeBottlePrimer207 : String;
      RPA30_scannedFrameBareCode : String;
      RPA30_Start : Bool;
      RPA30_cyclusState : UInt;
      RPA30_primer207_TimeExpiration : DTL;
      RPA30_Primer207_cycleCounter : Int;
      RPA30_stationState : Int;
      RPA30_ErrorStateLock : Int;
      RPA30_failStateLock : Int;
      RPA30_fatalErrorStateLock : Int;
      RPA30_bigFailStateLock : Int;
      RPA30_UseInterval_Primer207 : Bool;
      RPA30_valveYErrorStateCheck : Int;
      RPA30_scannedData : String;
      RPA30_bottle_taking : Bool;
      RPA30_UseIntervalBottleRemover208 : Bool;
      RPA30_actualCodeBottleRemover208 : String;
      RPA30_show_points_hmi : Byte;
   END_VAR
   VAR RETAIN
      RPA30_actual_instruction_index : Byte;
   END_VAR
   VAR
      RPA30_siren_hadler_enable : Bool;
      RPA30_pre_configuration : Byte;
   END_VAR
   VAR RETAIN
      RPA30_frame_581_Order : Int;
      RPA30_frame_582_Order : Int;
   END_VAR
   VAR
      RPA30_show_smile : Bool;
      RPA30_rotation_direction : Bool;
      RPA30_scaner_remover_counter : Byte;
      RPA30_remover_bottle_state_pre : Bool;
   END_VAR
   VAR RETAIN
      RPA30_station_configuration : Byte;
   END_VAR
   VAR
      RPA30_station_configuration_pre : Byte;
      RPA30_position_y_pre : Bool;
      RPA30_hmi_state_pre : Byte;
      RPA30_fail_state_pre : Int;
      RPA30_big_fail_state_pre : Int;
      RPA30_error_state_pre : Int;
      RPA30_fatal_error_state_pre : Int;
      RPA30_current_frame_code_pre : String;
      RPA30_state_information_send : Bool;
      RPA30_station_activity_state_pre : Bool;
      RPA30_show_pad_left : Bool;
      RPA30_show_pad_right : Bool;
      RPA30_side : Byte;
      RPA30_side_setup : Bool;
      RPA30_clock_pre : Bool;
      RPA30_rework_counter : UInt;
   END_VAR
   VAR RETAIN
      pa30_bottle_timing : LInt;
      pa30_bottle_cyclus_replace : UInt;
   END_VAR
   VAR
      pa30_left_ifm_connect_enable : Bool;
      pa30_right_ifm_connect_enable : Bool;
      pa30_right_ifm_change_application_enable : Bool;
      pa30_left_ifm_change_application_enable : Bool;
      pa30_left_ifm_application_index : UInt;
      pa30_right_ifm_application_index : UInt;
      pa30_right_ifm_actived_application_index : UInt;
      pa30_left_ifm_actived_application_index : UInt;
      pa30_right_ifm_data : Array[0..127] of Char;
      pa30_left_ifm_data : Array[0..127] of Char;
      pa30_left_size_in : UInt;
      pa30_right_size_in : UInt;
      pa30_right_status : UInt;
      pa30_left_status : UInt;
      pa30_done_left : Bool;
      pa30_done_right : Bool;
      pa30_ifm_triger_left : Bool;
      pa30_ifm_triger_right : Bool;
      pa30_ifm_left_busy : Bool;
      pa30_ifm_right_busy : Bool;
      pa30_ifm_right_error : Bool;
      pa30_ifm_left_error : Bool;
      pa30_keyence_switch : Bool;
      keyence_enable : Bool;
      ifm_run : Bool;
      ifm_side : Int;
   END_VAR
BEGIN
END_DATA_BLOCK

DATA_BLOCK "PA30_IFM_Left_PulsApplicationSwitch_DB"   // DB5
{ S7_Optimized_Access := 'FALSE' }
VERSION : 0.1
// stored: InstanceOfName IFM_PulsApplicationSwitch
"IFM_PulsApplicationSwitch"
BEGIN
END_DATA_BLOCK

DATA_BLOCK "PA30R_O2VxEth1500_left_DB"   // DB7
{ S7_Optimized_Access := 'FALSE' }
AUTHOR : ifm-sytl
FAMILY : O2Vx
NAME : O2Vx1500
VERSION : 1.3
// stored: InstanceOfName O2VxEth1500
"O2VxEth1500"
BEGIN
END_DATA_BLOCK

DATA_BLOCK "PLC_1_Send_DB"   // DB8
{ S7_Optimized_Access := 'FALSE' }
AUTHOR : SIMATIC
FAMILY : MC7Plus
NAME : TC_IP_v4
VERSION : 1.0
// stored: InstanceOfName ?
"?"
BEGIN
END_DATA_BLOCK

DATA_BLOCK "RPA30_F_TRIGR_DB"   // DB13
{ S7_Optimized_Access := 'FALSE' }
VERSION : 0.1
// stored: InstanceOfName RPA30_F_TRIGR
"RPA30_F_TRIGR"
BEGIN
END_DATA_BLOCK

DATA_BLOCK "print_label_PA60_DB"   // DB16
{ S7_Optimized_Access := 'FALSE' }
VERSION : 0.1
// stored: InstanceOfName print_label_PA60
"print_label_PA60"
BEGIN
END_DATA_BLOCK

DATA_BLOCK "PA10B_bottle_changing_DB"   // DB18
{ S7_Optimized_Access := 'FALSE' }
VERSION : 0.1
// stored: InstanceOfName bottle_changing
"bottle_changing"
BEGIN
END_DATA_BLOCK

DATA_BLOCK "RPA10B_datablock"   // DB19
{ S7_Optimized_Access := 'FALSE' }
VERSION : 0.1
   VAR
      PA10B_big_fail_state_lock : Int;
      PA10B_fail_state_lock : Int;
      PA10B_error_state_lock : Int;
      PA10B_fatal_error_state_lock : Int;
      RPA10B_station_start : Bool;
      PA10B_bottle_1_usage : Bool;
      PA10B_bottle_2_usage : Bool;
      PA10B_bottle_taking : Bool;
      RPA10B_station_work_cyclus_state : UInt;
      RPA10B_vacuum_activity_interval : UInt;
      RPA10B_idler_in_use : Bool;
      RPA10B_idler_taking : Bool;
      RPA10B_siren_hadler_enable : Bool;
      RPA10B_instruction_list_index : Byte;
      RPA10B_vacuum_R_check_state : Int;
      RPA10B_vacuum_L_check_state : Int;
      RPA10_valve_Y_check_state : Int;
      RPA10_valve_X_check_state : Int;
      RPA10B_end_of_cyclus : Bool;
      RPA10B_pad_checking_trigr : Bool;
      RPA10B_station_work_cyclus_state_pre : UInt;
      RPA10B_scanned_data : String;
      RPA10B_left_cover_code : String;
      RPA10B_right_cover_code : String;
      RPA10B_activator_bottle_1_code : String;
      RPA10B_activator_bottle_2_code : String;
      RPA10B_activator_bottle_1_cyclus_counter : Int;
      RPA10B_activator_bottle_1_expiration : DTL;
      RPA10B_activator_bottle_2_expiration : DTL;
      RPA10B_activator_bottle_2_cyclus_counter : Int;
      RPA10B_idler_checking_dalay : Bool;
      RPA10B_station_activity_state_pre : Bool;
      RPA10B_left_cover_code_pre : String;
      RPA10B_right_cover_code_pre : String;
      RPA10B_position_sensor_1_pre : Bool;
      RPA10B_position_sensor_2_pre : Bool;
      RPA10B_work_cyclus_state_pre : Byte;
      RPA10B_fail_state_pre : Int;
      RPA10B_big_fail_state_pre : Int;
      RPA10B_error_state_pre : Int;
      RPA10B_fata_error_state_pre : Int;
      RPA10B_station_monitoring_send : Bool;
      RPA10B_show_pad_left : Bool;
      RPA10B_show_pad_right : Bool;
      RPA10_B_show_home : Bool;
   END_VAR
   VAR RETAIN
      pa10B_bottle_timing : Time;
      pa10B_bottle_cyclus_replace : UInt;
   END_VAR
BEGIN
END_DATA_BLOCK

DATA_BLOCK "RPA20B_datablock"   // DB20
{ S7_Optimized_Access := 'FALSE' }
VERSION : 0.1
   VAR
      RPA20B_work_cyclus_state_OP_1 : Int;
      RPA20B_work_cyclus_state_OP_2 : Int;
      RPA20B_automatic_cyclus_enable : Bool;
      RPA20B_buffer_down_enable : Bool;
      RPA20B_activity_state_pre : Bool;
      RPA20B_left_cover_pressence_sensor_pre : Bool;
      RPA20B_right_cover_pressence_sensor_pre : Bool;
      RPA20B_station_monitoring_send : Bool;
   END_VAR
BEGIN
END_DATA_BLOCK

DATA_BLOCK "PA30_IFM_Right_PulsApplicationSwitch_DB"   // DB22
{ S7_Optimized_Access := 'FALSE' }
VERSION : 0.1
// stored: InstanceOfName IFM_PulsApplicationSwitch
"IFM_PulsApplicationSwitch"
BEGIN
END_DATA_BLOCK

DATA_BLOCK "RPA30_IFM_point_checking_DB"   // DB23
{ S7_Optimized_Access := 'FALSE' }
VERSION : 0.1
// stored: InstanceOfName PA30_IFM_point_checking
"PA30_IFM_point_checking"
BEGIN
END_DATA_BLOCK

DATA_BLOCK "PLC_datablock"   // DB26
{ S7_Optimized_Access := 'FALSE' }
VERSION : 0.1
   VAR RETAIN
      stations_configuration : Byte;
      frame_581_Order : Int;
      frame_582_Order : Int;
      frame_AU326_1_Order : Int;
   END_VAR
BEGIN
END_DATA_BLOCK

DATA_BLOCK "DB_RPA60_CAM"   // DB27
{ S7_Optimized_Access := 'FALSE' }
VERSION : 0.1
   VAR RETAIN
      RPA60_ENABLE_CAMERAS : Bool;
   END_VAR
BEGIN
END_DATA_BLOCK

DATA_BLOCK "RPA60_DataBlock"   // DB29
{ S7_Optimized_Access := 'FALSE' }
VERSION : 0.1
   VAR
      RPA60_valveYErrorStateCheck : Int;
      RPA60_fatalErrorStateLock : Int;
      RPA60_vacuumActivityInterval : UInt;
      RPA60_Start : Bool;
      RPA60_scannedFrameBareCode : String;
      RPA60_frameIndex : Int;
      RPA60_cyclusState : UInt;
      RPA60_ErrorStateLock : Int;
      RPA60_failStateLock : Int;
      RPA60_RollerDelay : Int;
      RPA60_rollerUsageInterval : Bool;
      RPA60_roller_taking : Bool;
      RPA60_bigFailStateLock : Int;
      RPA60_printEnable : Bool;
      RPA60_scanedData : String;
      RPA60_siren_hadler_enable : Bool;
      RPA60_hmi_instruction_index : Byte;
      RPA60_actual_time : DTL;
      RPA60_show_smile : Bool;
      RPA60_frame_order : String;
      RPA60_frame_record : Array[0..1023] of Char;
      RPA60_record_size : UInt;
      RPA60_station_configuration : Byte;
      RPA60_show_check_button : Bool;
      RPA60_number_of_check : Byte;
      RPA60_station_configuration_pre : Byte;
      RPA60_position_y_pre : Bool;
      RPA60_hmi_state_pre : Byte;
      RPA60_fail_state_pre : Int;
      RPA60_big_fail_state_pre : Int;
      RPA60_error_state_pre : Int;
      RPA60_fatal_error_state_pre : Int;
      RPA60_current_frame_code_pre : String;
      RPA60_state_information_send : Bool;
      RPA60_station_activity_state_pre : Bool;
      RPA60_rework_counter : UInt;
      RPA60_hardware_configuration : Byte;
      RPA60_side : Byte;
   END_VAR
BEGIN
END_DATA_BLOCK

DATA_BLOCK "PA10B_timer_lib_DB"   // DB30
{ S7_Optimized_Access := 'FALSE' }
VERSION : 0.1
// stored: InstanceOfName timer_lib
"timer_lib"
BEGIN
END_DATA_BLOCK

DATA_BLOCK "PA30R_O2VxEth1500_right_DB"   // DB31
{ S7_Optimized_Access := 'FALSE' }
AUTHOR : ifm-sytl
FAMILY : O2Vx
NAME : O2Vx1500
VERSION : 1.3
// stored: InstanceOfName O2VxEth1500
"O2VxEth1500"
BEGIN
END_DATA_BLOCK

DATA_BLOCK "PA30_timer_lib_DB"   // DB32
{ S7_Optimized_Access := 'FALSE' }
VERSION : 0.1
// stored: InstanceOfName timer_lib
"timer_lib"
BEGIN
END_DATA_BLOCK

DATA_BLOCK "pa60r_vacuum_cleaner_controll_DB"   // DB34
{ S7_Optimized_Access := 'FALSE' }
VERSION : 0.1
// stored: InstanceOfName vacuum_cleaner_controll
"vacuum_cleaner_controll"
BEGIN
END_DATA_BLOCK

DATA_BLOCK "TCP_Connection_DB"   // DB40
{ S7_Optimized_Access := 'FALSE' }
AUTHOR : SIMATIC
FAMILY : MC7Plus
NAME : TC_IP_v4
VERSION : 1.0
// stored: InstanceOfName ?
"?"
BEGIN
END_DATA_BLOCK

DATA_BLOCK "PA60R_timer_lib_DB"   // DB45
{ S7_Optimized_Access := 'FALSE' }
VERSION : 0.1
// stored: InstanceOfName timer_lib
"timer_lib"
BEGIN
END_DATA_BLOCK

DATA_BLOCK "fs_print_label_fce_DB"   // DB46
{ S7_Optimized_Access := 'FALSE' }
VERSION : 0.1
// stored: InstanceOfName fs_print_label_fce
"fs_print_label_fce"
BEGIN
END_DATA_BLOCK

DATA_BLOCK "tcp_datablock"   // DB48
{ S7_Optimized_Access := 'FALSE' }
VERSION : 0.1
   VAR
      index_send : Byte;
      index_out : Byte;
      tcp_connection : Bool;
      "counter" : UInt;
      ping_index : Byte;
      fs_shaker_1_index : Byte;
      fs_shaker_2_index : Byte;
      fs_shaker_3_index : Byte;
      fs_shaker_4_index : Byte;
      fs_shaker_5_index : Byte;
      fs_fill_bottle_index : Byte;
      pa10b_handler_index : Byte;
      pa60r_station_state_index : Byte;
      pa20b_station_state_index : Byte;
      pa10b_station_state_index : Byte;
      pa30r_station_state_index : Byte;
      pa60r_handler_index : Byte;
      pa30r_handler_index : Byte;
      fs_print_sp_label_index : Byte;
      tcp_size_out : Array[0..5] of UInt;
      tcp_transaction_done : Array[0..5] of Bool;
      tcp_input_buffer : Array[0..5] of "tcp_data_item";
      tcp_output_buffer : Array[0..5] of "tcp_data_item";
   END_VAR
BEGIN
END_DATA_BLOCK

DATA_BLOCK "pa10b_vacuum_cleaner_controll_DB"   // DB49
{ S7_Optimized_Access := 'FALSE' }
VERSION : 0.1
// stored: InstanceOfName vacuum_cleaner_controll
"vacuum_cleaner_controll"
BEGIN
END_DATA_BLOCK

// folder: System blocks/Program resources

DATA_BLOCK "IEC_Timer_0_DB"   // DB6
{ S7_Optimized_Access := 'FALSE' }
AUTHOR : Simatic
FAMILY : IEC
NAME : IEC_TMR
VERSION : 1.0
// stored: InstanceOfName ?
"?"
BEGIN
END_DATA_BLOCK

DATA_BLOCK "PA20B_Timer_0_DB"   // DB37
{ S7_Optimized_Access := 'FALSE' }
AUTHOR : Simatic
FAMILY : IEC
NAME : IEC_TMR
VERSION : 1.0
// stored: InstanceOfName ?
"?"
BEGIN
END_DATA_BLOCK

DATA_BLOCK "PA20B_Timer_1_DB"   // DB39
{ S7_Optimized_Access := 'FALSE' }
AUTHOR : Simatic
FAMILY : IEC
NAME : IEC_TMR
VERSION : 1.0
// stored: InstanceOfName ?
"?"
BEGIN
END_DATA_BLOCK

DATA_BLOCK "printer_connection"   // DB43
{ S7_Optimized_Access := 'FALSE' }
AUTHOR : SIMATIC
FAMILY : MC7Plus
NAME : TC_IP_v4
VERSION : 1.0
// stored: InstanceOfName ?
"?"
BEGIN
END_DATA_BLOCK

// folder: (top level)

FUNCTION_BLOCK "IFM_PulsApplicationSwitch"   // FB1, SCL
{ S7_Optimized_Access := 'FALSE' }
VERSION : 0.1
BEGIN
   IF #IFM_switch_enable THEN
       IF #IFM_ApplicationIndex > 0 THEN
           CASE #IFM_Switch_State OF
               0:
                   #IFM_Application_Switched := false;
                   #IFM_Input_1 := true;
                   #IFM_Pulse_Number := #IFM_ApplicationIndex;
                   //change the state to the next value
                   #IFM_Switch_State := 1;
               1:
                   //pulsing in precisely time intervals
                   #timer_lib_Instance(#IFM_Pulse_Period);
                   IF #IFM_Pulse_Number > 0 THEN
                       IF #IFM_Input_2 = false AND #timer_lib_Instance.DONE THEN
                           #IFM_Input_2 := true;
                       ELSIF #IFM_Input_2 = true AND #timer_lib_Instance.DONE THEN
                           #IFM_Pulse_Number := #IFM_Pulse_Number - 1;
                           #IFM_Input_2 := false;
                       END_IF;
                   ELSE
                       // set input 1 to false
                       #IFM_Input_1 := false;
                       #IFM_Switch_State := 2;

                   END_IF;
               2:
                   IF #ready_intput = false THEN
                       #IFM_Switch_State := 3;
                   END_IF;

               3:
                   #timer_lib_Instance(3000);
                   IF #timer_lib_Instance.DONE THEN
                       #IFM_Switch_State := 0;
                       #timer_lib_Instance.lock := false;
                   END_IF;

                   IF #ready_intput = true THEN
                       #IFM_Switch_State := 0;
                       //set free to switch of application       
                       #IFM_Application_Switched := true;
                       #IFM_switch_enable := false;
                       #timer_lib_Instance.lock := false;
                   END_IF;

               ELSE  // Statement section ELSE
                   #IFM_Switch_State := 0;
                   #IFM_Input_1 := false;
                   #IFM_Input_2 := false;
                    #IFM_Application_Switched := false;
                   #IFM_switch_enable :=false;
           END_CASE;
       END_IF;
   END_IF;

   (*

   IF #IFM_ApplicationIndex > 0 THEN
       CASE #IFM_Application_Switch_State OF
           0: //set state switching of application

               #IFM_Input_1 := true;
               //change the state to the next value